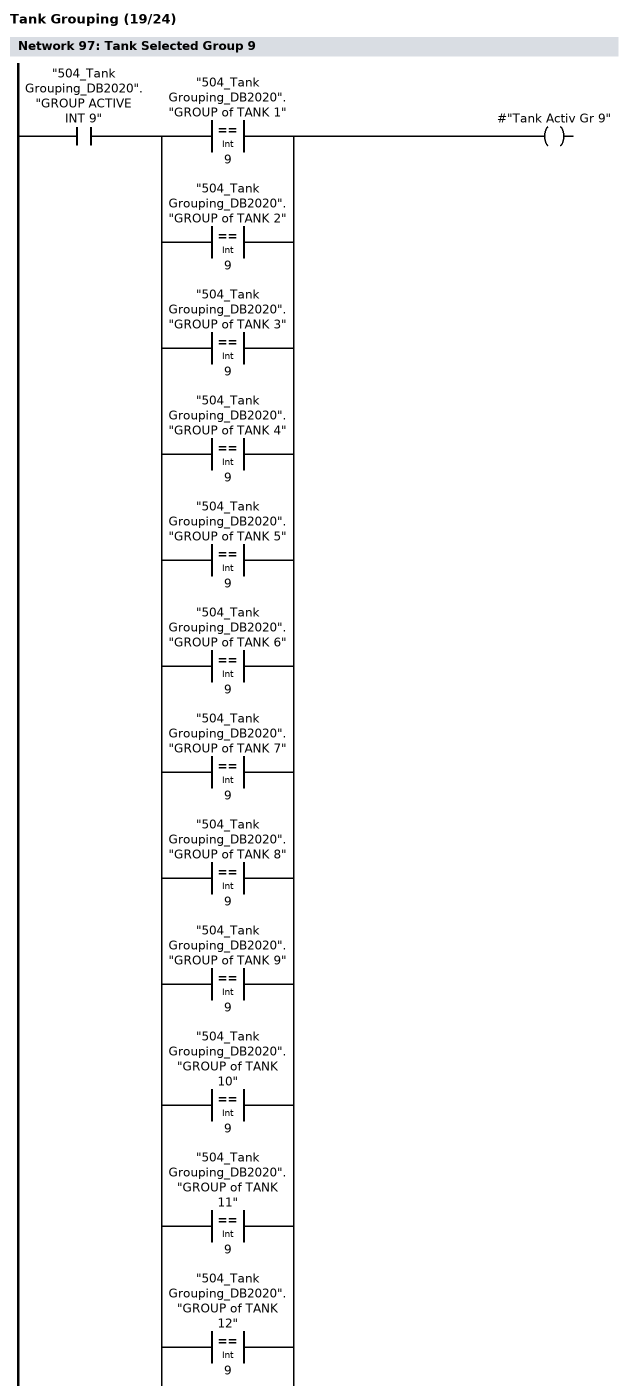
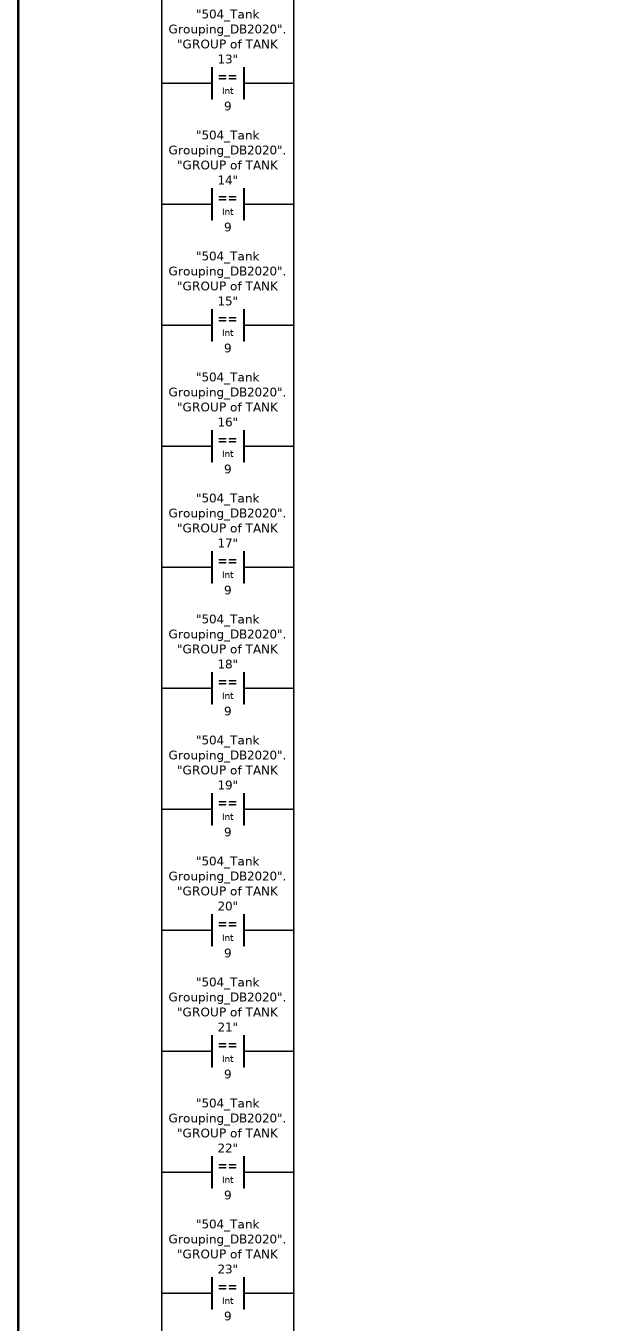
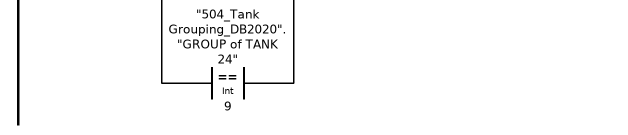
   RUNG wire#powerrail
      Contact( "504_Tank Grouping_DB2020"."GROUP ACTIVE INT 9" )
      wire#w1
      { S7_Templates := "SrcType := Int" } EQ_Contact(in1 := "504_Tank Grouping_DB2020"."GROUP of TANK 1", in2 := 9)
      wire#w2
      Coil( #"Tank Activ Gr 9" )
   END_RUNG
   RUNG wire#w1
      { S7_Templates := "SrcType := Int" } EQ_Contact(in1 := "504_Tank Grouping_DB2020"."GROUP of TANK 2", in2 := 9)
   END_RUNG wire#w2
   RUNG wire#w1
      { S7_Templates := "SrcType := Int" } EQ_Contact(in1 := "504_Tank Grouping_DB2020"."GROUP of TANK 3", in2 := 9)
   END_RUNG wire#w2
   RUNG wire#w1
      { S7_Templates := "SrcType := Int" } EQ_Contact(in1 := "504_Tank Grouping_DB2020"."GROUP of TANK 4", in2 := 9)
   END_RUNG wire#w2
   RUNG wire#w1
      { S7_Templates := "SrcType := Int" } EQ_Contact(in1 := "504_Tank Grouping_DB2020"."GROUP of TANK 5", in2 := 9)
   END_RUNG wire#w2
   RUNG wire#w1
      { S7_Templates := "SrcType := Int" } EQ_Contact(in1 := "504_Tank Grouping_DB2020"."GROUP of TANK 6", in2 := 9)
   END_RUNG wire#w2
   RUNG wire#w1
      { S7_Templates := "SrcType := Int" } EQ_Contact(in1 := "504_Tank Grouping_DB2020"."GROUP of TANK 7", in2 := 9)
   END_RUNG wire#w2
   RUNG wire#w1
      { S7_Templates := "SrcType := Int" } EQ_Contact(in1 := "504_Tank Grouping_DB2020"."GROUP of TANK 8", in2 := 9)
   END_RUNG wire#w2
   RUNG wire#w1
      { S7_Templates := "SrcType := Int" } EQ_Contact(in1 := "504_Tank Grouping_DB2020"."GROUP of TANK 9", in2 := 9)
   END_RUNG wire#w2
   RUNG wire#w1
      { S7_Templates := "SrcType := Int" } EQ_Contact(in1 := "504_Tank Grouping_DB2020"."GROUP of TANK 10", in2 := 9)
   END_RUNG wire#w2
   RUNG wire#w1
      { S7_Templates := "SrcType := Int" } EQ_Contact(in1 := "504_Tank Grouping_DB2020"."GROUP of TANK 11", in2 := 9)
   END_RUNG wire#w2
   RUNG wire#w1
      { S7_Templates := "SrcType := Int" } EQ_Contact(in1 := "504_Tank Grouping_DB2020"."GROUP of TANK 12", in2 := 9)
   END_RUNG wire#w2
   RUNG wire#w1
      { S7_Templates := "SrcType := Int" } EQ_Contact(in1 := "504_Tank Grouping_DB2020"."GROUP of TANK 13", in2 := 9)
   END_RUNG wire#w2
   RUNG wire#w1
      { S7_Templates := "SrcType := Int" } EQ_Contact(in1 := "504_Tank Grouping_DB2020"."GROUP of TANK 14", in2 := 9)
   END_RUNG wire#w2
   RUNG wire#w1
      { S7_Templates := "SrcType := Int" } EQ_Contact(in1 := "504_Tank Grouping_DB2020"."GROUP of TANK 15", in2 := 9)
   END_RUNG wire#w2
   RUNG wire#w1
      { S7_Templates := "SrcType := Int" } EQ_Contact(in1 := "504_Tank Grouping_DB2020"."GROUP of TANK 16", in2 := 9)
   END_RUNG wire#w2
   RUNG wire#w1
      { S7_Templates := "SrcType := Int" } EQ_Contact(in1 := "504_Tank Grouping_DB2020"."GROUP of TANK 17", in2 := 9)
   END_RUNG wire#w2
   RUNG wire#w1
      { S7_Templates := "SrcType := Int" } EQ_Contact(in1 := "504_Tank Grouping_DB2020"."GROUP of TANK 18", in2 := 9)
   END_RUNG wire#w2
   RUNG wire#w1
      { S7_Templates := "SrcType := Int" } EQ_Contact(in1 := "504_Tank Grouping_DB2020"."GROUP of TANK 19", in2 := 9)
   END_RUNG wire#w2
   RUNG wire#w1
      { S7_Templates := "SrcType := Int" } EQ_Contact(in1 := "504_Tank Grouping_DB2020"."GROUP of TANK 20", in2 := 9)
   END_RUNG wire#w2
   RUNG wire#w1
      { S7_Templates := "SrcType := Int" } EQ_Contact(in1 := "504_Tank Grouping_DB2020"."GROUP of TANK 21", in2 := 9)
   END_RUNG wire#w2
   RUNG wire#w1
      { S7_Templates := "SrcType := Int" } EQ_Contact(in1 := "504_Tank Grouping_DB2020"."GROUP of TANK 22", in2 := 9)
   END_RUNG wire#w2
   RUNG wire#w1
      { S7_Templates := "SrcType := Int" } EQ_Contact(in1 := "504_Tank Grouping_DB2020"."GROUP of TANK 23", in2 := 9)
   END_RUNG wire#w2
   RUNG wire#w1
      { S7_Templates := "SrcType := Int" } EQ_Contact(in1 := "504_Tank Grouping_DB2020"."GROUP of TANK 24", in2 := 9)
   END_RUNG wire#w2
   // the same network as SCL:
   #"Tank Activ Gr 9" := "504_Tank Grouping_DB2020"."GROUP ACTIVE INT 9" AND (("504_Tank Grouping_DB2020"."GROUP of TANK 1" = 9) OR ("504_Tank Grouping_DB2020"."GROUP of TANK 2" = 9) OR ("504_Tank Grouping_DB2020"."GROUP of TANK 3" = 9) OR ("504_Tank Grouping_DB2020"."GROUP of TANK 4" = 9) OR ("504_Tank Grouping_DB2020"."GROUP of TANK 5" = 9) OR ("504_Tank Grouping_DB2020"."GROUP of TANK 6" = 9) OR ("504_Tank Grouping_DB2020"."GROUP of TANK 7" = 9) OR ("504_Tank Grouping_DB2020"."GROUP of TANK 8" = 9) OR ("504_Tank Grouping_DB2020"."GROUP of TANK 9" = 9) OR ("504_Tank Grouping_DB2020"."GROUP of TANK 10" = 9) OR ("504_Tank Grouping_DB2020"."GROUP of TANK 11" = 9) OR ("504_Tank Grouping_DB2020"."GROUP of TANK 12" = 9) OR ("504_Tank Grouping_DB2020"."GROUP of TANK 13" = 9) OR ("504_Tank Grouping_DB2020"."GROUP of TANK 14" = 9) OR ("504_Tank Grouping_DB2020"."GROUP of TANK 15" = 9) OR ("504_Tank Grouping_DB2020"."GROUP of TANK 16" = 9) OR ("504_Tank Grouping_DB2020"."GROUP of TANK 17" = 9) OR ("504_Tank Grouping_DB2020"."GROUP of TANK 18" = 9) OR ("504_Tank Grouping_DB2020"."GROUP of TANK 19" = 9) OR ("504_Tank Grouping_DB2020"."GROUP of TANK 20" = 9) OR ("504_Tank Grouping_DB2020"."GROUP of TANK 21" = 9) OR ("504_Tank Grouping_DB2020"."GROUP of TANK 22" = 9) OR ("504_Tank Grouping_DB2020"."GROUP of TANK 23" = 9) OR ("504_Tank Grouping_DB2020"."GROUP of TANK 24" = 9));
END_REGION

REGION Network 98: Tank Selected Group 10
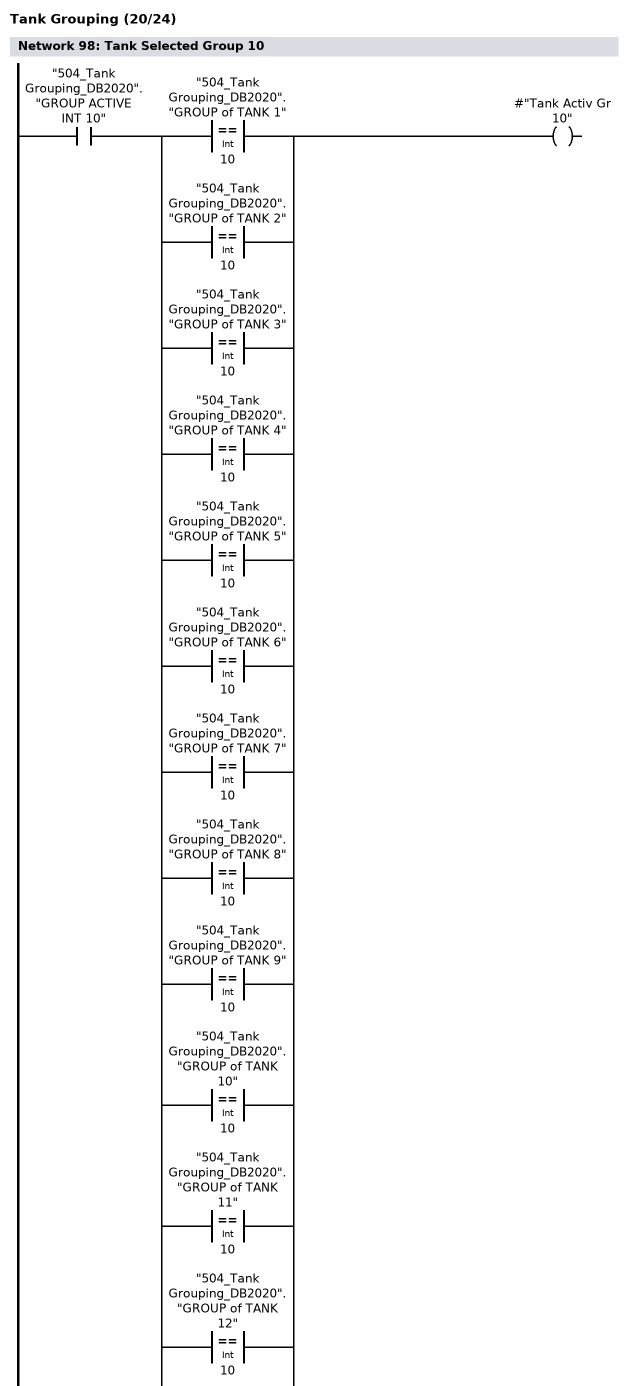
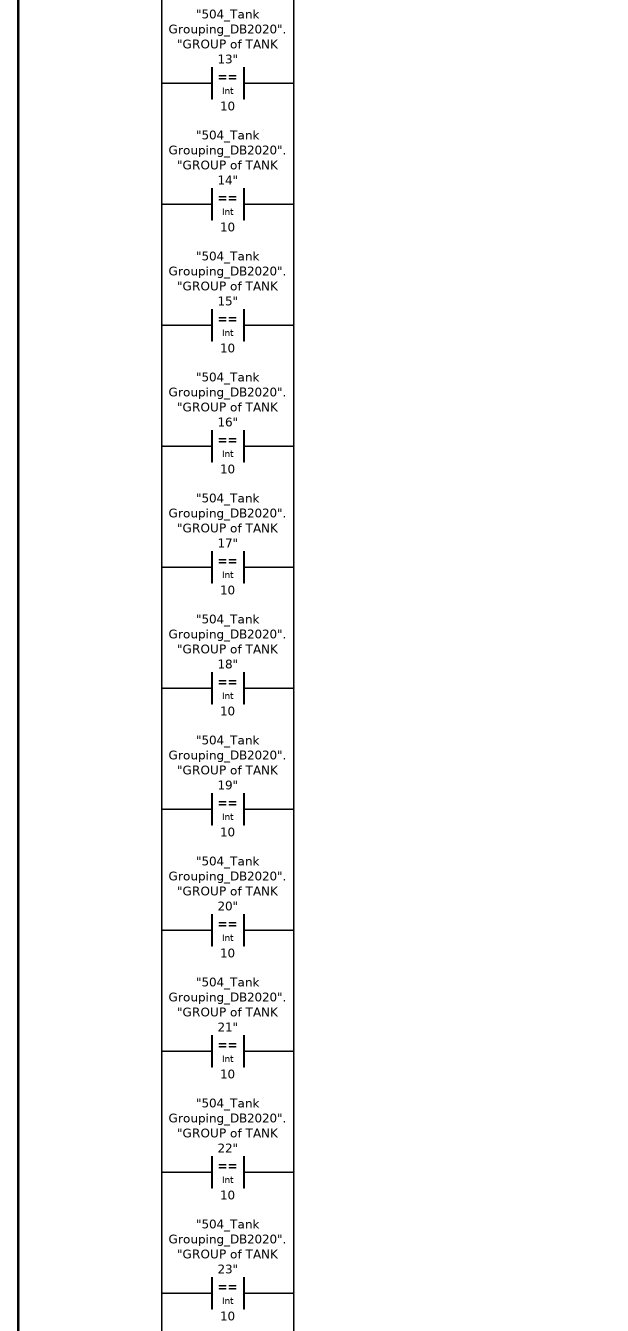
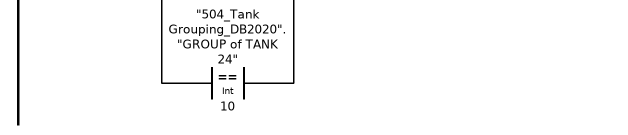
   RUNG wire#powerrail
      Contact( "504_Tank Grouping_DB2020"."GROUP ACTIVE INT 10" )
      wire#w1
      { S7_Templates := "SrcType := Int" } EQ_Contact(in1 := "504_Tank Grouping_DB2020"."GROUP of TANK 1", in2 := 10)
      wire#w2
      Coil( #"Tank Activ Gr 10" )
   END_RUNG
   RUNG wire#w1
      { S7_Templates := "SrcType := Int" } EQ_Contact(in1 := "504_Tank Grouping_DB2020"."GROUP of TANK 2", in2 := 10)
   END_RUNG wire#w2
   RUNG wire#w1
      { S7_Templates := "SrcType := Int" } EQ_Contact(in1 := "504_Tank Grouping_DB2020"."GROUP of TANK 3", in2 := 10)
   END_RUNG wire#w2
   RUNG wire#w1
      { S7_Templates := "SrcType := Int" } EQ_Contact(in1 := "504_Tank Grouping_DB2020"."GROUP of TANK 4", in2 := 10)
   END_RUNG wire#w2
   RUNG wire#w1
      { S7_Templates := "SrcType := Int" } EQ_Contact(in1 := "504_Tank Grouping_DB2020"."GROUP of TANK 5", in2 := 10)
   END_RUNG wire#w2
   RUNG wire#w1
      { S7_Templates := "SrcType := Int" } EQ_Contact(in1 := "504_Tank Grouping_DB2020"."GROUP of TANK 6", in2 := 10)
   END_RUNG wire#w2
   RUNG wire#w1
      { S7_Templates := "SrcType := Int" } EQ_Contact(in1 := "504_Tank Grouping_DB2020"."GROUP of TANK 7", in2 := 10)
   END_RUNG wire#w2
   RUNG wire#w1
      { S7_Templates := "SrcType := Int" } EQ_Contact(in1 := "504_Tank Grouping_DB2020"."GROUP of TANK 8", in2 := 10)
   END_RUNG wire#w2
   RUNG wire#w1
      { S7_Templates := "SrcType := Int" } EQ_Contact(in1 := "504_Tank Grouping_DB2020"."GROUP of TANK 9", in2 := 10)
   END_RUNG wire#w2
   RUNG wire#w1
      { S7_Templates := "SrcType := Int" } EQ_Contact(in1 := "504_Tank Grouping_DB2020"."GROUP of TANK 10", in2 := 10)
   END_RUNG wire#w2
   RUNG wire#w1
      { S7_Templates := "SrcType := Int" } EQ_Contact(in1 := "504_Tank Grouping_DB2020"."GROUP of TANK 11", in2 := 10)
   END_RUNG wire#w2
   RUNG wire#w1
      { S7_Templates := "SrcType := Int" } EQ_Contact(in1 := "504_Tank Grouping_DB2020"."GROUP of TANK 12", in2 := 10)
   END_RUNG wire#w2
   RUNG wire#w1
      { S7_Templates := "SrcType := Int" } EQ_Contact(in1 := "504_Tank Grouping_DB2020"."GROUP of TANK 13", in2 := 10)
   END_RUNG wire#w2
   RUNG wire#w1
      { S7_Templates := "SrcType := Int" } EQ_Contact(in1 := "504_Tank Grouping_DB2020"."GROUP of TANK 14", in2 := 10)
   END_RUNG wire#w2
   RUNG wire#w1
      { S7_Templates := "SrcType := Int" } EQ_Contact(in1 := "504_Tank Grouping_DB2020"."GROUP of TANK 15", in2 := 10)
   END_RUNG wire#w2
   RUNG wire#w1
      { S7_Templates := "SrcType := Int" } EQ_Contact(in1 := "504_Tank Grouping_DB2020"."GROUP of TANK 16", in2 := 10)
   END_RUNG wire#w2
   RUNG wire#w1
      { S7_Templates := "SrcType := Int" } EQ_Contact(in1 := "504_Tank Grouping_DB2020"."GROUP of TANK 17", in2 := 10)
   END_RUNG wire#w2
   RUNG wire#w1
      { S7_Templates := "SrcType := Int" } EQ_Contact(in1 := "504_Tank Grouping_DB2020"."GROUP of TANK 18", in2 := 10)
   END_RUNG wire#w2
   RUNG wire#w1
      { S7_Templates := "SrcType := Int" } EQ_Contact(in1 := "504_Tank Grouping_DB2020"."GROUP of TANK 19", in2 := 10)
   END_RUNG wire#w2
   RUNG wire#w1
      { S7_Templates := "SrcType := Int" } EQ_Contact(in1 := "504_Tank Grouping_DB2020"."GROUP of TANK 20", in2 := 10)
   END_RUNG wire#w2
   RUNG wire#w1
      { S7_Templates := "SrcType := Int" } EQ_Contact(in1 := "504_Tank Grouping_DB2020"."GROUP of TANK 21", in2 := 10)
   END_RUNG wire#w2
   RUNG wire#w1
      { S7_Templates := "SrcType := Int" } EQ_Contact(in1 := "504_Tank Grouping_DB2020"."GROUP of TANK 22", in2 := 10)
   END_RUNG wire#w2
   RUNG wire#w1
      { S7_Templates := "SrcType := Int" } EQ_Contact(in1 := "504_Tank Grouping_DB2020"."GROUP of TANK 23", in2 := 10)
   END_RUNG wire#w2
   RUNG wire#w1
      { S7_Templates := "SrcType := Int" } EQ_Contact(in1 := "504_Tank Grouping_DB2020"."GROUP of TANK 24", in2 := 10)
   END_RUNG wire#w2
   // the same network as SCL:
   #"Tank Activ Gr 10" := "504_Tank Grouping_DB2020"."GROUP ACTIVE INT 10" AND (("504_Tank Grouping_DB2020"."GROUP of TANK 1" = 10) OR ("504_Tank Grouping_DB2020"."GROUP of TANK 2" = 10) OR ("504_Tank Grouping_DB2020"."GROUP of TANK 3" = 10) OR ("504_Tank Grouping_DB2020"."GROUP of TANK 4" = 10) OR ("504_Tank Grouping_DB2020"."GROUP of TANK 5" = 10) OR ("504_Tank Grouping_DB2020"."GROUP of TANK 6" = 10) OR ("504_Tank Grouping_DB2020"."GROUP of TANK 7" = 10) OR ("504_Tank Grouping_DB2020"."GROUP of TANK 8" = 10) OR ("504_Tank Grouping_DB2020"."GROUP of TANK 9" = 10) OR ("504_Tank Grouping_DB2020"."GROUP of TANK 10" = 10) OR ("504_Tank Grouping_DB2020"."GROUP of TANK 11" = 10) OR ("504_Tank Grouping_DB2020"."GROUP of TANK 12" = 10) OR ("504_Tank Grouping_DB2020"."GROUP of TANK 13" = 10) OR ("504_Tank Grouping_DB2020"."GROUP of TANK 14" = 10) OR ("504_Tank Grouping_DB2020"."GROUP of TANK 15" = 10) OR ("504_Tank Grouping_DB2020"."GROUP of TANK 16" = 10) OR ("504_Tank Grouping_DB2020"."GROUP of TANK 17" = 10) OR ("504_Tank Grouping_DB2020"."GROUP of TANK 18" = 10) OR ("504_Tank Grouping_DB2020"."GROUP of TANK 19" = 10) OR ("504_Tank Grouping_DB2020"."GROUP of TANK 20" = 10) OR ("504_Tank Grouping_DB2020"."GROUP of TANK 21" = 10) OR ("504_Tank Grouping_DB2020"."GROUP of TANK 22" = 10) OR ("504_Tank Grouping_DB2020"."GROUP of TANK 23" = 10) OR ("504_Tank Grouping_DB2020"."GROUP of TANK 24" = 10));
END_REGION

REGION Network 99: Tank Selected Group 12
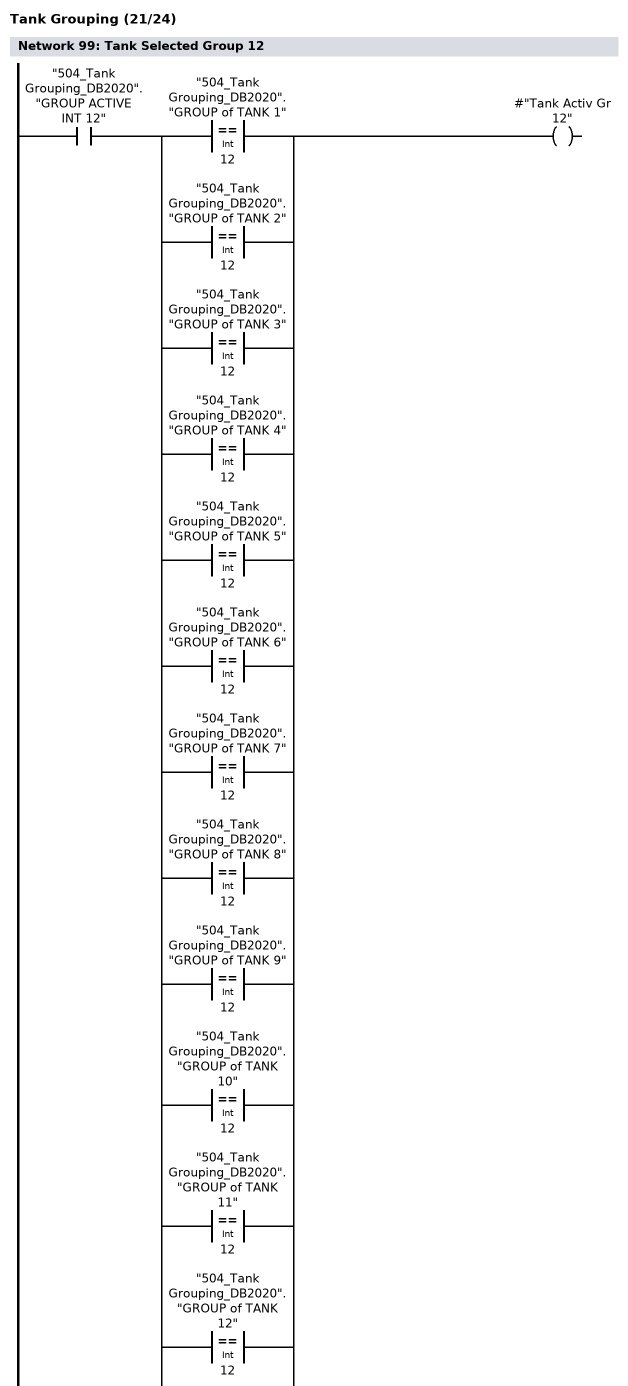
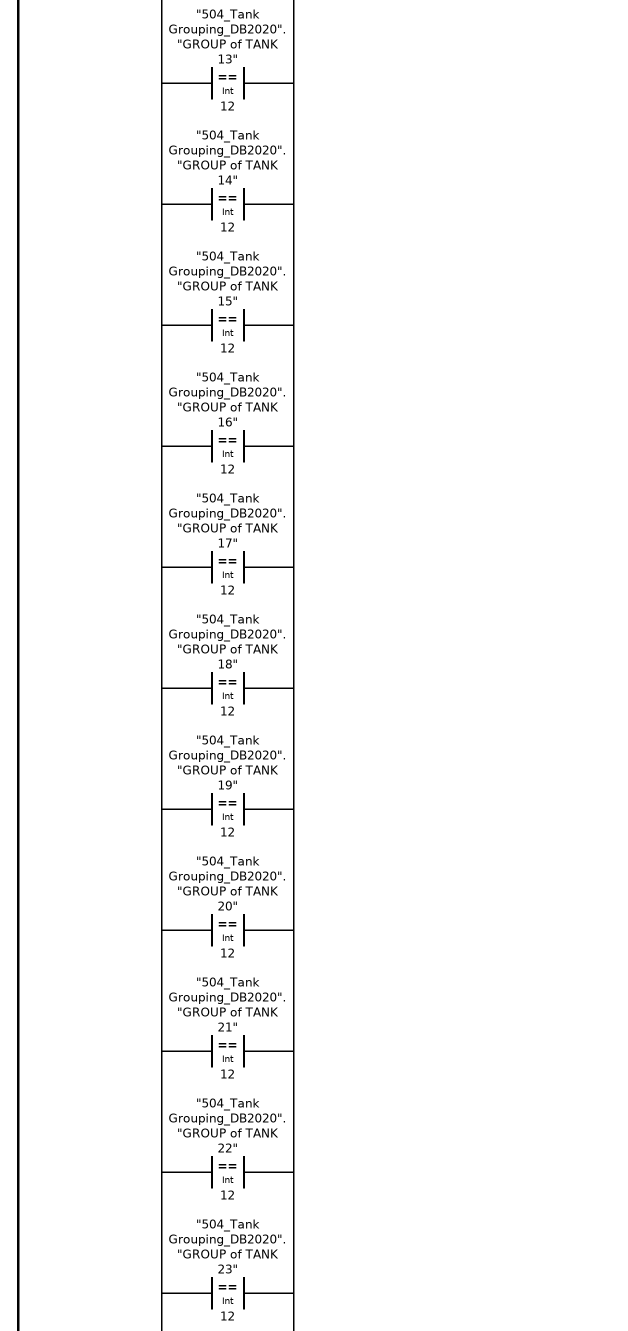
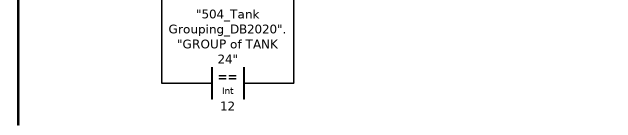
   RUNG wire#powerrail
      Contact( "504_Tank Grouping_DB2020"."GROUP ACTIVE INT 12" )
      wire#w1
      { S7_Templates := "SrcType := Int" } EQ_Contact(in1 := "504_Tank Grouping_DB2020"."GROUP of TANK 1", in2 := 12)
      wire#w2
      Coil( #"Tank Activ Gr 12" )
   END_RUNG
   RUNG wire#w1
      { S7_Templates := "SrcType := Int" } EQ_Contact(in1 := "504_Tank Grouping_DB2020"."GROUP of TANK 2", in2 := 12)
   END_RUNG wire#w2
   RUNG wire#w1
      { S7_Templates := "SrcType := Int" } EQ_Contact(in1 := "504_Tank Grouping_DB2020"."GROUP of TANK 3", in2 := 12)
   END_RUNG wire#w2
   RUNG wire#w1
      { S7_Templates := "SrcType := Int" } EQ_Contact(in1 := "504_Tank Grouping_DB2020"."GROUP of TANK 4", in2 := 12)
   END_RUNG wire#w2
   RUNG wire#w1
      { S7_Templates := "SrcType := Int" } EQ_Contact(in1 := "504_Tank Grouping_DB2020"."GROUP of TANK 5", in2 := 12)
   END_RUNG wire#w2
   RUNG wire#w1
      { S7_Templates := "SrcType := Int" } EQ_Contact(in1 := "504_Tank Grouping_DB2020"."GROUP of TANK 6", in2 := 12)
   END_RUNG wire#w2
   RUNG wire#w1
      { S7_Templates := "SrcType := Int" } EQ_Contact(in1 := "504_Tank Grouping_DB2020"."GROUP of TANK 7", in2 := 12)
   END_RUNG wire#w2
   RUNG wire#w1
      { S7_Templates := "SrcType := Int" } EQ_Contact(in1 := "504_Tank Grouping_DB2020"."GROUP of TANK 8", in2 := 12)
   END_RUNG wire#w2
   RUNG wire#w1
      { S7_Templates := "SrcType := Int" } EQ_Contact(in1 := "504_Tank Grouping_DB2020"."GROUP of TANK 9", in2 := 12)
   END_RUNG wire#w2
   RUNG wire#w1
      { S7_Templates := "SrcType := Int" } EQ_Contact(in1 := "504_Tank Grouping_DB2020"."GROUP of TANK 10", in2 := 12)
   END_RUNG wire#w2
   RUNG wire#w1
      { S7_Templates := "SrcType := Int" } EQ_Contact(in1 := "504_Tank Grouping_DB2020"."GROUP of TANK 11", in2 := 12)
   END_RUNG wire#w2
   RUNG wire#w1
      { S7_Templates := "SrcType := Int" } EQ_Contact(in1 := "504_Tank Grouping_DB2020"."GROUP of TANK 12", in2 := 12)
   END_RUNG wire#w2
   RUNG wire#w1
      { S7_Templates := "SrcType := Int" } EQ_Contact(in1 := "504_Tank Grouping_DB2020"."GROUP of TANK 13", in2 := 12)
   END_RUNG wire#w2
   RUNG wire#w1
      { S7_Templates := "SrcType := Int" } EQ_Contact(in1 := "504_Tank Grouping_DB2020"."GROUP of TANK 14", in2 := 12)
   END_RUNG wire#w2
   RUNG wire#w1
      { S7_Templates := "SrcType := Int" } EQ_Contact(in1 := "504_Tank Grouping_DB2020"."GROUP of TANK 15", in2 := 12)
   END_RUNG wire#w2
   RUNG wire#w1
      { S7_Templates := "SrcType := Int" } EQ_Contact(in1 := "504_Tank Grouping_DB2020"."GROUP of TANK 16", in2 := 12)
   END_RUNG wire#w2
   RUNG wire#w1
      { S7_Templates := "SrcType := Int" } EQ_Contact(in1 := "504_Tank Grouping_DB2020"."GROUP of TANK 17", in2 := 12)
   END_RUNG wire#w2
   RUNG wire#w1
      { S7_Templates := "SrcType := Int" } EQ_Contact(in1 := "504_Tank Grouping_DB2020"."GROUP of TANK 18", in2 := 12)
   END_RUNG wire#w2
   RUNG wire#w1
      { S7_Templates := "SrcType := Int" } EQ_Contact(in1 := "504_Tank Grouping_DB2020"."GROUP of TANK 19", in2 := 12)
   END_RUNG wire#w2
   RUNG wire#w1
      { S7_Templates := "SrcType := Int" } EQ_Contact(in1 := "504_Tank Grouping_DB2020"."GROUP of TANK 20", in2 := 12)
   END_RUNG wire#w2
   RUNG wire#w1
      { S7_Templates := "SrcType := Int" } EQ_Contact(in1 := "504_Tank Grouping_DB2020"."GROUP of TANK 21", in2 := 12)
   END_RUNG wire#w2
   RUNG wire#w1
      { S7_Templates := "SrcType := Int" } EQ_Contact(in1 := "504_Tank Grouping_DB2020"."GROUP of TANK 22", in2 := 12)
   END_RUNG wire#w2
   RUNG wire#w1
      { S7_Templates := "SrcType := Int" } EQ_Contact(in1 := "504_Tank Grouping_DB2020"."GROUP of TANK 23", in2 := 12)
   END_RUNG wire#w2
   RUNG wire#w1
      { S7_Templates := "SrcType := Int" } EQ_Contact(in1 := "504_Tank Grouping_DB2020"."GROUP of TANK 24", in2 := 12)
   END_RUNG wire#w2
   // the same network as SCL:
   #"Tank Activ Gr 12" := "504_Tank Grouping_DB2020"."GROUP ACTIVE INT 12" AND (("504_Tank Grouping_DB2020"."GROUP of TANK 1" = 12) OR ("504_Tank Grouping_DB2020"."GROUP of TANK 2" = 12) OR ("504_Tank Grouping_DB2020"."GROUP of TANK 3" = 12) OR ("504_Tank Grouping_DB2020"."GROUP of TANK 4" = 12) OR ("504_Tank Grouping_DB2020"."GROUP of TANK 5" = 12) OR ("504_Tank Grouping_DB2020"."GROUP of TANK 6" = 12) OR ("504_Tank Grouping_DB2020"."GROUP of TANK 7" = 12) OR ("504_Tank Grouping_DB2020"."GROUP of TANK 8" = 12) OR ("504_Tank Grouping_DB2020"."GROUP of TANK 9" = 12) OR ("504_Tank Grouping_DB2020"."GROUP of TANK 10" = 12) OR ("504_Tank Grouping_DB2020"."GROUP of TANK 11" = 12) OR ("504_Tank Grouping_DB2020"."GROUP of TANK 12" = 12) OR ("504_Tank Grouping_DB2020"."GROUP of TANK 13" = 12) OR ("504_Tank Grouping_DB2020"."GROUP of TANK 14" = 12) OR ("504_Tank Grouping_DB2020"."GROUP of TANK 15" = 12) OR ("504_Tank Grouping_DB2020"."GROUP of TANK 16" = 12) OR ("504_Tank Grouping_DB2020"."GROUP of TANK 17" = 12) OR ("504_Tank Grouping_DB2020"."GROUP of TANK 18" = 12) OR ("504_Tank Grouping_DB2020"."GROUP of TANK 19" = 12) OR ("504_Tank Grouping_DB2020"."GROUP of TANK 20" = 12) OR ("504_Tank Grouping_DB2020"."GROUP of TANK 21" = 12) OR ("504_Tank Grouping_DB2020"."GROUP of TANK 22" = 12) OR ("504_Tank Grouping_DB2020"."GROUP of TANK 23" = 12) OR ("504_Tank Grouping_DB2020"."GROUP of TANK 24" = 12));
END_REGION

REGION Network 100: Tank Selected Group 13
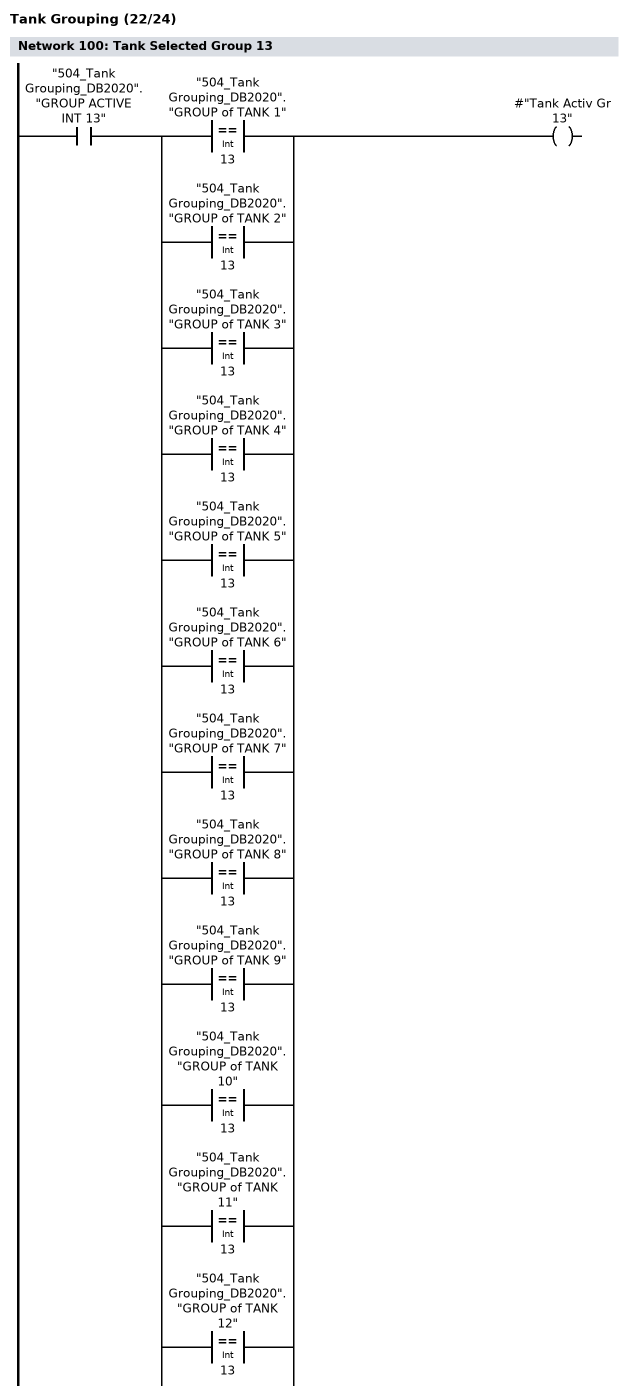
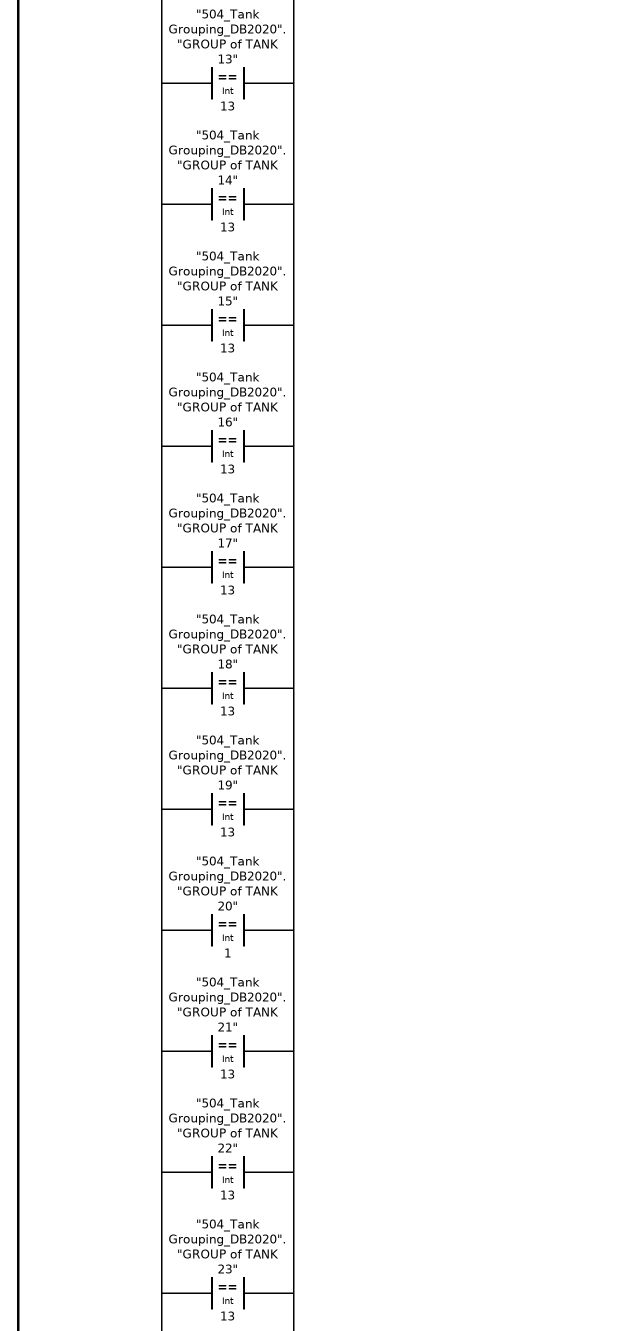
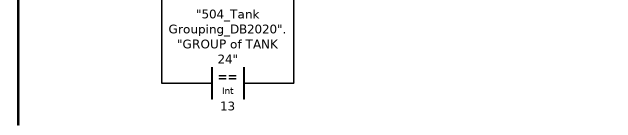
   RUNG wire#powerrail
      Contact( "504_Tank Grouping_DB2020"."GROUP ACTIVE INT 13" )
      wire#w1
      { S7_Templates := "SrcType := Int" } EQ_Contact(in1 := "504_Tank Grouping_DB2020"."GROUP of TANK 1", in2 := 13)
      wire#w2
      Coil( #"Tank Activ Gr 13" )
   END_RUNG
   RUNG wire#w1
      { S7_Templates := "SrcType := Int" } EQ_Contact(in1 := "504_Tank Grouping_DB2020"."GROUP of TANK 2", in2 := 13)
   END_RUNG wire#w2
   RUNG wire#w1
      { S7_Templates := "SrcType := Int" } EQ_Contact(in1 := "504_Tank Grouping_DB2020"."GROUP of TANK 3", in2 := 13)
   END_RUNG wire#w2
   RUNG wire#w1
      { S7_Templates := "SrcType := Int" } EQ_Contact(in1 := "504_Tank Grouping_DB2020"."GROUP of TANK 4", in2 := 13)
   END_RUNG wire#w2
   RUNG wire#w1
      { S7_Templates := "SrcType := Int" } EQ_Contact(in1 := "504_Tank Grouping_DB2020"."GROUP of TANK 5", in2 := 13)
   END_RUNG wire#w2
   RUNG wire#w1
      { S7_Templates := "SrcType := Int" } EQ_Contact(in1 := "504_Tank Grouping_DB2020"."GROUP of TANK 6", in2 := 13)
   END_RUNG wire#w2
   RUNG wire#w1
      { S7_Templates := "SrcType := Int" } EQ_Contact(in1 := "504_Tank Grouping_DB2020"."GROUP of TANK 7", in2 := 13)
   END_RUNG wire#w2
   RUNG wire#w1
      { S7_Templates := "SrcType := Int" } EQ_Contact(in1 := "504_Tank Grouping_DB2020"."GROUP of TANK 8", in2 := 13)
   END_RUNG wire#w2
   RUNG wire#w1
      { S7_Templates := "SrcType := Int" } EQ_Contact(in1 := "504_Tank Grouping_DB2020"."GROUP of TANK 9", in2 := 13)
   END_RUNG wire#w2
   RUNG wire#w1
      { S7_Templates := "SrcType := Int" } EQ_Contact(in1 := "504_Tank Grouping_DB2020"."GROUP of TANK 10", in2 := 13)
   END_RUNG wire#w2
   RUNG wire#w1
      { S7_Templates := "SrcType := Int" } EQ_Contact(in1 := "504_Tank Grouping_DB2020"."GROUP of TANK 11", in2 := 13)
   END_RUNG wire#w2
   RUNG wire#w1
      { S7_Templates := "SrcType := Int" } EQ_Contact(in1 := "504_Tank Grouping_DB2020"."GROUP of TANK 12", in2 := 13)
   END_RUNG wire#w2
   RUNG wire#w1
      { S7_Templates := "SrcType := Int" } EQ_Contact(in1 := "504_Tank Grouping_DB2020"."GROUP of TANK 13", in2 := 13)
   END_RUNG wire#w2
   RUNG wire#w1
      { S7_Templates := "SrcType := Int" } EQ_Contact(in1 := "504_Tank Grouping_DB2020"."GROUP of TANK 14", in2 := 13)
   END_RUNG wire#w2
   RUNG wire#w1
      { S7_Templates := "SrcType := Int" } EQ_Contact(in1 := "504_Tank Grouping_DB2020"."GROUP of TANK 15", in2 := 13)
   END_RUNG wire#w2
   RUNG wire#w1
      { S7_Templates := "SrcType := Int" } EQ_Contact(in1 := "504_Tank Grouping_DB2020"."GROUP of TANK 16", in2 := 13)
   END_RUNG wire#w2
   RUNG wire#w1
      { S7_Templates := "SrcType := Int" } EQ_Contact(in1 := "504_Tank Grouping_DB2020"."GROUP of TANK 17", in2 := 13)
   END_RUNG wire#w2
   RUNG wire#w1
      { S7_Templates := "SrcType := Int" } EQ_Contact(in1 := "504_Tank Grouping_DB2020"."GROUP of TANK 18", in2 := 13)
   END_RUNG wire#w2
   RUNG wire#w1
      { S7_Templates := "SrcType := Int" } EQ_Contact(in1 := "504_Tank Grouping_DB2020"."GROUP of TANK 19", in2 := 13)
   END_RUNG wire#w2
   RUNG wire#w1
      { S7_Templates := "SrcType := Int" } EQ_Contact(in1 := "504_Tank Grouping_DB2020"."GROUP of TANK 20", in2 := 1)
   END_RUNG wire#w2
   RUNG wire#w1
      { S7_Templates := "SrcType := Int" } EQ_Contact(in1 := "504_Tank Grouping_DB2020"."GROUP of TANK 21", in2 := 13)
   END_RUNG wire#w2
   RUNG wire#w1
      { S7_Templates := "SrcType := Int" } EQ_Contact(in1 := "504_Tank Grouping_DB2020"."GROUP of TANK 22", in2 := 13)
   END_RUNG wire#w2
   RUNG wire#w1
      { S7_Templates := "SrcType := Int" } EQ_Contact(in1 := "504_Tank Grouping_DB2020"."GROUP of TANK 23", in2 := 13)
   END_RUNG wire#w2
   RUNG wire#w1
      { S7_Templates := "SrcType := Int" } EQ_Contact(in1 := "504_Tank Grouping_DB2020"."GROUP of TANK 24", in2 := 13)
   END_RUNG wire#w2
   // the same network as SCL:
   #"Tank Activ Gr 13" := "504_Tank Grouping_DB2020"."GROUP ACTIVE INT 13" AND (("504_Tank Grouping_DB2020"."GROUP of TANK 1" = 13) OR ("504_Tank Grouping_DB2020"."GROUP of TANK 2" = 13) OR ("504_Tank Grouping_DB2020"."GROUP of TANK 3" = 13) OR ("504_Tank Grouping_DB2020"."GROUP of TANK 4" = 13) OR ("504_Tank Grouping_DB2020"."GROUP of TANK 5" = 13) OR ("504_Tank Grouping_DB2020"."GROUP of TANK 6" = 13) OR ("504_Tank Grouping_DB2020"."GROUP of TANK 7" = 13) OR ("504_Tank Grouping_DB2020"."GROUP of TANK 8" = 13) OR ("504_Tank Grouping_DB2020"."GROUP of TANK 9" = 13) OR ("504_Tank Grouping_DB2020"."GROUP of TANK 10" = 13) OR ("504_Tank Grouping_DB2020"."GROUP of TANK 11" = 13) OR ("504_Tank Grouping_DB2020"."GROUP of TANK 12" = 13) OR ("504_Tank Grouping_DB2020"."GROUP of TANK 13" = 13) OR ("504_Tank Grouping_DB2020"."GROUP of TANK 14" = 13) OR ("504_Tank Grouping_DB2020"."GROUP of TANK 15" = 13) OR ("504_Tank Grouping_DB2020"."GROUP of TANK 16" = 13) OR ("504_Tank Grouping_DB2020"."GROUP of TANK 17" = 13) OR ("504_Tank Grouping_DB2020"."GROUP of TANK 18" = 13) OR ("504_Tank Grouping_DB2020"."GROUP of TANK 19" = 13) OR ("504_Tank Grouping_DB2020"."GROUP of TANK 20" = 1) OR ("504_Tank Grouping_DB2020"."GROUP of TANK 21" = 13) OR ("504_Tank Grouping_DB2020"."GROUP of TANK 22" = 13) OR ("504_Tank Grouping_DB2020"."GROUP of TANK 23" = 13) OR ("504_Tank Grouping_DB2020"."GROUP of TANK 24" = 13));
END_REGION

REGION Network 101: Tank Selected Group 14
